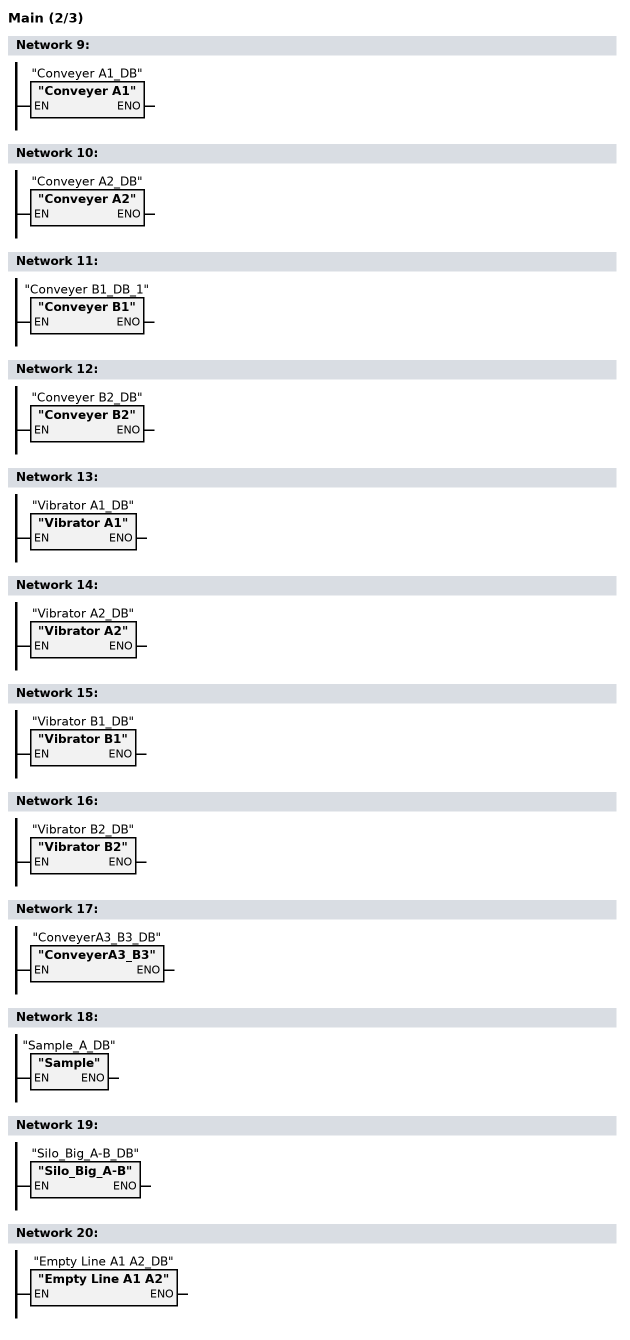
   RUNG wire#powerrail
      "Conveyer A1_DB"()
   END_RUNG
   // the same network as SCL:
   "Conveyer A1_DB"();   // "Conveyer A1"
END_REGION

REGION Network 10
   RUNG wire#powerrail
      "Conveyer A2_DB"()
   END_RUNG
   // the same network as SCL:
   "Conveyer A2_DB"();   // "Conveyer A2"
END_REGION

REGION Network 11
   RUNG wire#powerrail
      "Conveyer B1_DB_1"()
   END_RUNG
   // the same network as SCL:
   "Conveyer B1_DB_1"();   // "Conveyer B1"
END_REGION

REGION Network 12
   RUNG wire#powerrail
      "Conveyer B2_DB"()
   END_RUNG
   // the same network as SCL:
   "Conveyer B2_DB"();   // "Conveyer B2"
END_REGION

REGION Network 13
   RUNG wire#powerrail
      "Vibrator A1_DB"()
   END_RUNG
   // the same network as SCL:
   "Vibrator A1_DB"();   // "Vibrator A1"
END_REGION

REGION Network 14
   RUNG wire#powerrail
      "Vibrator A2_DB"()
   END_RUNG
   // the same network as SCL:
   "Vibrator A2_DB"();   // "Vibrator A2"
END_REGION

REGION Network 15
   RUNG wire#powerrail
      "Vibrator B1_DB"()
   END_RUNG
   // the same network as SCL:
   "Vibrator B1_DB"();   // "Vibrator B1"
END_REGION

REGION Network 16
   RUNG wire#powerrail
      "Vibrator B2_DB"()
   END_RUNG
   // the same network as SCL:
   "Vibrator B2_DB"();   // "Vibrator B2"
END_REGION

REGION Network 17
   RUNG wire#powerrail
      "ConveyerA3_B3_DB"()
   END_RUNG
   // the same network as SCL:
   "ConveyerA3_B3_DB"();   // "ConveyerA3_B3"
END_REGION

REGION Network 18
   RUNG wire#powerrail
      "Sample_A_DB"()
   END_RUNG
   // the same network as SCL:
   "Sample_A_DB"();   // "Sample"
END_REGION

REGION Network 19
   RUNG wire#powerrail
      "Silo_Big_A-B_DB"()
   END_RUNG
   // the same network as SCL:
   "Silo_Big_A-B_DB"();   // "Silo_Big_A-B"
END_REGION

REGION Network 20
   RUNG wire#powerrail
      "Empty Line A1 A2_DB"()
   END_RUNG
   // the same network as SCL:
   "Empty Line A1 A2_DB"();   // "Empty Line A1 A2"
END_REGION

REGION Network 21
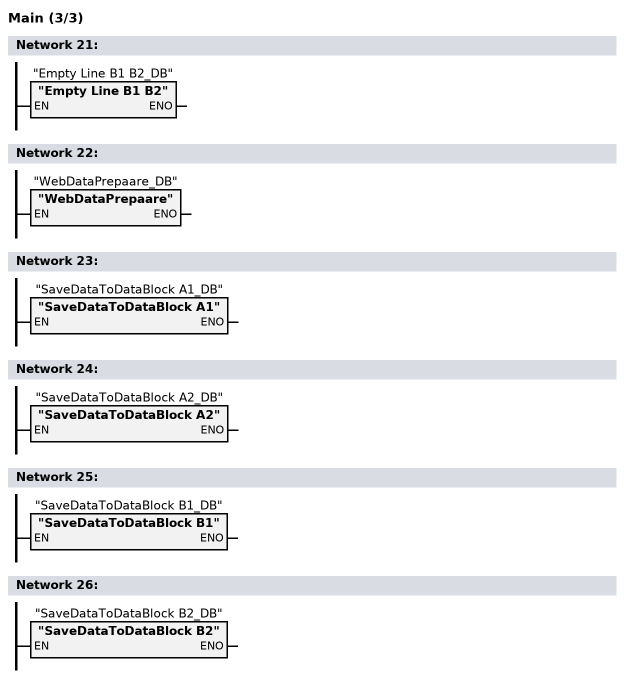
   RUNG wire#powerrail
      "Empty Line B1 B2_DB"()
   END_RUNG
   // the same network as SCL:
   "Empty Line B1 B2_DB"();   // "Empty Line B1 B2"
END_REGION

REGION Network 22
   RUNG wire#powerrail
      "WebDataPrepaare_DB"()
   END_RUNG
   // the same network as SCL:
   "WebDataPrepaare_DB"();   // "WebDataPrepaare"
END_REGION

REGION Network 23
   RUNG wire#powerrail
      "SaveDataToDataBlock A1_DB"()
   END_RUNG
   // the same network as SCL:
   "SaveDataToDataBlock A1_DB"();   // "SaveDataToDataBlock A1"
END_REGION

REGION Network 24
   RUNG wire#powerrail
      "SaveDataToDataBlock A2_DB"()
   END_RUNG
   // the same network as SCL:
   "SaveDataToDataBlock A2_DB"();   // "SaveDataToDataBlock A2"
END_REGION

REGION Network 25
   RUNG wire#powerrail
      "SaveDataToDataBlock B1_DB"()
   END_RUNG
   // the same network as SCL:
   "SaveDataToDataBlock B1_DB"();   // "SaveDataToDataBlock B1"
END_REGION

REGION Network 26
   RUNG wire#powerrail
      "SaveDataToDataBlock B2_DB"()
   END_RUNG
   // the same network as SCL:
   "SaveDataToDataBlock B2_DB"();   // "SaveDataToDataBlock B2"
END_REGION
END_ORGANIZATION_BLOCK

// ===== PLC "PLC_Lines_C"  CPU 1212C AC/DC/Rly =====

VAR_GLOBAL   // PLC tag table "Default tag table"
   "Tag_4" AT %MW114 : Word;
   "Tag_5" AT %M118.0 : Bool;
   "Tag_6" AT %M118.1 : Bool;
   "Tag_7" AT %M118.2 : Bool;
   "Tag_8" AT %MW120 : Word;
   "Tag_9" AT %MW122 : Word;
   "Tag_1" AT %M251.0 : Bool;
   "C2_Start_Conveyer" AT %M161.1 : Bool;
   "Tag_3" AT %M1000.0 : Bool;
   "Tag_10" AT %M1200.0 : Bool;
   "Vibrator_C1_On" AT %M151.4 : Bool;
   "Tag_11" AT %M151.5 : Bool;
   "Tag_2" AT %M123.2 : Bool;
   "Vibrator_C2_On" AT %M161.4 : Bool;
   "Tag_12" AT %M160.6 : Bool;
   "Conveyer_C2_On" AT %M160.3 : Bool;
   "Tag_13" AT %M161.5 : Bool;
   "Tag_14" AT %M151.7 : Bool;
   "Conveyer_C1_OneShut" AT %M151.3 : Bool;
   "Conveyer_C2_OneShut" AT %M161.3 : Bool;
   "Silo C Big" AT %Q3.6 : Bool;
   "Silo_C_Big_Start_Toggle" AT %M190.0 : Bool;
   "TriggerStartToggleMemory" AT %M152.0 : Bool;
   "TriggerC1ToggleStop" AT %M152.1 : Bool;
   "Conveyor_C1_Empty_line" AT %M152.2 : Bool;
   "Line_C2_Conveyer_Timer" AT %M162.0 : Bool;
   "TriggerStartToggleMemoryC2" AT %M162.1 : Bool;
   "TriggerStopToggleMemoryC21" AT %M162.2 : Bool;
   "Conveyor_C2_Empty_line" AT %M162.3 : Bool;
   "Silo_C_Not_Start_Timer" AT %M180.0 : Bool;
   "SiloCToggleStart" AT %M180.1 : Bool;
   "Tag_15" AT %MD210 : DInt;
   "Tag_16" AT %MD240 : DInt;
   "Tag_17" AT %M500.1 : Bool;
   "Tag_18" AT %M500.2 : Bool;
   "Tag_24" AT %MW502 : Word;
   "Tag_26" AT %M504.0 : Bool;
   "Tag_27" AT %M504.1 : Bool;
   "Tag_28" AT %M504.2 : Bool;
   "Tag_29" AT %MW506 : Word;
   "Tag_30" AT %MW508 : Word;
   "Tag_31" AT %MW510 : Word;
   "Tag_32" AT %M504.7 : Bool;
END_VAR

VAR_GLOBAL   // PLC tag table "InputOutput"
   "Emergency_C" AT %I0.6 : Bool;   // OK
   "Low_Silo_C1" AT %I0.2 : Bool;   // OK
   "Conveyer_C1" AT %Q0.2 : Bool;   // OK
   "Conveyer_C2" AT %Q0.3 : Bool;   // OK
   "Rel Out Vibrator C1" AT %Q0.0 : Bool;
   "Rel Out Vibrator C2" AT %Q0.1 : Bool;
   "Rel Out Alarm C1" AT %Q2.2 : Bool;
   "Rel Out Alarm C2" AT %Q2.3 : Bool;
   "Pneumatic_C1" AT %Q0.4 : Bool;   // OK
   "Pneumatic_C2" AT %Q0.5 : Bool;   // OK
   "Rel Out Conveyer C" AT %Q2.4 : Bool;
   "Rel Out Silo C Stop" AT %Q2.5 : Bool;
   "Rel Out Silo C Start" AT %Q2.6 : Bool;
   "Low_Silo_C2" AT %I0.0 : Bool;   // OK
   "HIgh_Silo_C1" AT %I0.3 : Bool;   // OK
   "Fault_C1" AT %I0.4 : Bool;   // OK
   "Fault_C2" AT %I0.5 : Bool;   // OK
   "High_Silo_C2" AT %I0.1 : Bool;   // OK
   "Start" AT %I1.1 : Bool;
   "Fault_C3" AT %I0.7 : Bool;   // OK
   "Conveyer_C3" AT %Q3.4 : Bool;   // OK
   "Light_C1" AT %Q2.0 : Bool;   // OK
   "Light_C2" AT %Q2.1 : Bool;   // OK
END_VAR

VAR_GLOBAL   // PLC tag table "SystemTag"
   "System_Byte" AT %MB1 : Byte;
   "FirstScan" AT %M1.0 : Bool;
   "DiagStatusUpdate" AT %M1.1 : Bool;
   "AlwaysTRUE" AT %M1.2 : Bool;
   "AlwaysFALSE" AT %M1.3 : Bool;
   "Clock_Byte" AT %MB0 : Byte;
   "Clock_10Hz" AT %M0.0 : Bool;
   "Clock_5Hz" AT %M0.1 : Bool;
   "Clock_2.5Hz" AT %M0.2 : Bool;
   "Clock_2Hz" AT %M0.3 : Bool;
   "Clock_1.25Hz" AT %M0.4 : Bool;
   "Clock_1Hz" AT %M0.5 : Bool;
   "Clock_0.625Hz" AT %M0.6 : Bool;
   "Clock_0.5Hz" AT %M0.7 : Bool;
   "DoneModbusCommon" AT %M110.0 : Bool;
   "ErrorModbusCommon" AT %M110.1 : Bool;
   "ModbusCommonStatus" AT %MW112 : Word;
END_VAR

VAR_GLOBAL   // PLC tag table "LineC1Tags"
   "Line_C1_Start_Consent" AT %M150.0 : Bool;
   "Line_C1_Run_Consent" AT %M150.1 : Bool;
   "Line_C1_Conveyer_Timer" AT %M150.2 : Bool;
   "Conveyer_C1_On" AT %M150.3 : Bool;
   "Conveyer_C1_Off" AT %M150.4 : Bool;
   "Line_C1_Light" AT %M151.0 : Bool;
   "Start_C1_Toggle" AT %M150.5 : Bool;
   "StartTriggerRisingTrigger" AT %M150.6 : Bool;
   "Conveyer_C1_Start_Consent" AT %M250.0 : Bool;
   "Conveyer_C1_Run_Consent" AT %M250.1 : Bool;
   "Silo_C_Start" AT %M300.0 : Bool;
   "C1_Sample_Triger" AT %M150.7 : Bool;
   "C1_Start_Conveyer" AT %M151.1 : Bool;
END_VAR

VAR_GLOBAL   // PLC tag table "LineC2Tags"
   "Line_C2_Start_Consent" AT %M160.0 : Bool;
   "Line_C2_Run_Consent" AT %M160.1 : Bool;
   "Line_C2_Vibrator_Timer" AT %M160.2 : Bool;
   "Conveyer_C2_Off" AT %M160.4 : Bool;
   "Conveyer_C2_Start_Consent" AT %M260.0 : Bool;
   "Conveyer_C2_Run_Consent" AT %M260.1 : Bool;
   "Start_C2_Toggle" AT %M160.5 : Bool;
   "C2_Sample_Triger" AT %M160.7 : Bool;
END_VAR

TYPE "tIMEDATATYPE"
   STRUCT
      HOUR : String;
      MINUTE : String;
      DAY : String;
      MONTH : String;
      YEAR : String;
   END_STRUCT;
END_TYPE

DATA_BLOCK "ModbusDataSendToFeeders"   // DB7
{ S7_Optimized_Access := 'FALSE' }
VERSION : 0.1
   VAR
      dataforsend : Array[0..3] of Int;
   END_VAR
BEGIN
   dataforsend[0] := 0;
   dataforsend[1] := 0;
   dataforsend[2] := 0;
   dataforsend[3] := 0;
END_DATA_BLOCK

DATA_BLOCK "Clock"   // DB9
{ S7_Optimized_Access := 'TRUE' }
VERSION : 0.1
   VAR
      "time" : DTL;
   END_VAR
BEGIN
END_DATA_BLOCK

DATA_BLOCK "Conveyer C1_DB"   // DB16
{ S7_Optimized_Access := 'TRUE' }
VERSION : 0.1
// stored: InstanceOfName Conveyer C1
"Conveyer C1"
BEGIN
END_DATA_BLOCK

DATA_BLOCK "Web_Send"   // DB23
{ S7_Optimized_Access := 'TRUE' }
VERSION : 0.1
   VAR
      C1_Scenario_Type : Int := 2;
      C2_Scenario_Type : Int := 1;
      B1_Scenario_Type : Int := 1;
      B2_Scenario_Type : Int := 1;
      C_Emergency : Bool;
      B_Emergency : Bool;
      C1_Fault : Bool;
      C2_Fault : Bool;
      B1_Fault : Bool;
      B2_Fault : Bool;
      C3_Fault : Bool;
      B3_Fault : Bool;
      C1_Silo_Low : Bool;
      C2_Silo_Low : Bool;
      B1_Silo_Low : Bool;
      B2_Silo_Low : Bool;
      C1_Conveyer : Bool;
      C2_Conveyer : Bool;
      B1_Conveyer : Bool;
      B2_Conveyer : Bool;
      C3_Conveyor : Bool;
      B3_Left_Conveyer : Bool;
      C1_Silo_High : Bool;
      C2_Silo_High : Bool;
      B1_Silo_High : Bool;
      B2_Silo_High : Bool;
      C1_Sample : Bool;
      C2_Sample : Bool;
      B1_Sample : Bool;
      B2_Sample : Bool;
      C1_Running_Duration : Time;
      C1_Pause_Duration : Time;
      C1_Feeder_Vibration_Intensity : Int;
      C1_Ruuning_Online : Time;
      C1_Pause_Online : Time;
      C1_Sample_Interval : Time;
      C1_Sample_Duration : Time;
      C1_Sample_Online : Time;
      C1_Enable : Bool;
      C1_Start : Bool;
      C1_Big_Silo : Bool;
      B1_Running_Duration : Time;
      B1_Pause_Duration : Time;
      B1_Feeder_Vibration_Intensity : Int;
      B1_Ruuning_Online : Time;
      B1_Pause_Online : Time;
      B1_Sample_Interval : Time;
      B1_Sample_Duration : Time;
      B1_Sample_Online : Time;
      B1_Enable : Bool;
      B1_Start : Bool;
      B1_Big_Silo : Bool;
      C2_Running_Duration : Time;
      C2_Pause_Duration : Time;
      C2_Feeder_Vibration_Intensity : Int;
      C2_Ruuning_Online : Time;
      C2_Pause_Online : Time;
      C2_Sample_Interval : Time;
      C2_Sample_Duration : Time;
      C2_Sample_Online : Time;
      C2_Enable : Bool;
      C2_Start : Bool;
      C2_Big_Silo : Bool;
      B2_Running_Duration : Time;
      B2_Pause_Duration : Time;
      B2_Feeder_Vibration_Intensity : Int;
      B2_Ruuning_Online : Time;
      B2_Pause_Online : Time;
      B2_Sample_Interval : Time;
      B2_Sample_Duration : Time;
      B2_Sample_Online : Time;
      B2_Enable : Bool;
      B2_Start : Bool;
      B2_Big_Silo : Bool;
      C1_Manual : Bool;
      C2_Manual : Bool;
      B1_Manual : Bool;
      B2_Manual : Bool;
      C1_Feeder : Bool;
      C2_Feeder : Bool;
      B1_Feeder : Bool;
      B2_Feeder : Bool;
      C1_Duration_Big_Silo_Stop_Time : Time;
      C2_Duration_Big_Silo_Stop_Time : Time;
      B1_Duration_Big_Silo_Stop_Time : Time;
      B2_Duration_Big_Silo_Stop_Time : Time;
      C1_Empty_Line_Time : Time;
      C2_Empty_Line_Time : Time;
      B1_Empty_Line_Time : Time;
      B2_Empty_Line_Time : Time;
      C1_Feeder_Delay_After_Start_Time : Time;
      C2_Feeder_Delay_After_Start_Time : Time;
      B1_Feeder_Delay_After_Start_Time : Time;
      B2_Feeder_Delay_After_Start_Time : Time;
      C1_Feeder_Delay_Before_Stop_Time : Time;
      C2_Feeder_Delay_Before_Stop_Time : Time;
      B1_Feeder_Delay_Before_Stop_Time : Time;
      B2_Feeder_Delay_Before_Stop_Time : Time;
      C1_Feeder_Delay_Time : Time;
      C1_Feeder_Delay_Time_1 : Time;
      C1_Feeder_Delay_Time_2 : Time;
      C1_Feeder_Delay_Time_3 : Time;
      B3_Conveyor : Bool;
   END_VAR
BEGIN
END_DATA_BLOCK

DATA_BLOCK "Conveyer C2_DB"   // DB24
{ S7_Optimized_Access := 'TRUE' }
VERSION : 0.1
// stored: InstanceOfName Conveyer C2
"Conveyer C2"
BEGIN
END_DATA_BLOCK

DATA_BLOCK "Vibrator C1_DB"   // DB25
{ S7_Optimized_Access := 'TRUE' }
VERSION : 0.1
// stored: InstanceOfName Vibrator C1
"Vibrator C1"
BEGIN
END_DATA_BLOCK

DATA_BLOCK "Vibrator C2_DB"   // DB26
{ S7_Optimized_Access := 'TRUE' }
VERSION : 0.1
// stored: InstanceOfName Vibrator C2
"Vibrator C2"
BEGIN
END_DATA_BLOCK

DATA_BLOCK "ConveyerC3_DB"   // DB35
{ S7_Optimized_Access := 'TRUE' }
VERSION : 0.1
// stored: InstanceOfName ConveyerC3
"ConveyerC3"
BEGIN
END_DATA_BLOCK

DATA_BLOCK "Sample_C_DB"   // DB36
{ S7_Optimized_Access := 'TRUE' }
VERSION : 0.1
// stored: InstanceOfName Sample_C
"Sample_C"
BEGIN
END_DATA_BLOCK

DATA_BLOCK "Silo_Big_C_DB"   // DB37
{ S7_Optimized_Access := 'TRUE' }
VERSION : 0.1
// stored: InstanceOfName Silo_Big_C
"Silo_Big_C"
BEGIN
END_DATA_BLOCK

DATA_BLOCK "Empty Line C1_DB"   // DB38
{ S7_Optimized_Access := 'TRUE' }
VERSION : 0.1
// stored: InstanceOfName Empty Line C1
"Empty Line C1"
BEGIN
END_DATA_BLOCK

DATA_BLOCK "Web_Recieve"   // DB45
{ S7_Optimized_Access := 'TRUE' }
VERSION : 0.1
   VAR
      Scenario_Type : Int;   // 1 2 3 4 5 A B C D E F
      Line_C1_Start : Bool;
      Line_C1_Enable : Bool := 0;
      Line_C2_Start : Bool;
      Line_C2_Enable : Bool;
      Line_C1_Conveyer_on_Time : Time := T#8S_400MS;
      Line_C1_Conveyer_off_Time : Time := T#30s;
      Line_C1_Sampling_Time : Time := T#2M;
      Line_C1_Sampling_OpenTime : Time := T#9S_500MS;
      Line_C2_Conveyer_on_Time : Time := T#8S_400MS;
      Line_C2_Conveyer_off_Time : Time := T#30s;
      Line_C2_Sampling_Time : Time := T#2M;
      Line_C2_Sampling_OpenTime : Time := T#9S_500MS;
      Line_C1_Feeder_Intensity : Int;
      Line_C2_Feeder_Intensity : Int;
      Line_C1_Feeder_DelayTime : Time;
      Line_C2_Feeder_DelayTime : Time;
      Line_C1_Enable_Manual : Bool;
      Line_C2_Enable_Manual : Bool;
      Line_C1_Conveyor_Start_Manual : Bool;
      Line_C2_Conveyor_Start_Manual : Bool;
      Line_C1_Big_Silo_Start_Manual : Bool;
      Line_C2_Big_Silo_Start_Manual : Bool;
      Line_C1_Below_Conveyor_Start_Manual : Bool;
      Line_C2_Below_Conveyor_Start_Manual : Bool;
      Line_C1_Feeder_Start_Manual : Bool;
      Line_C2_Feeder_Start_Manual : Bool;
      Line_B1_Feeder_Start_Manual : Bool;
      Line_B2_Feeder_Start_Manual : Bool;
      Line_C1_Sample_Start_Manual : Bool;
      Line_C2_Sample_Start_Manual : Bool;
      Line_B1_Sample_Start_Manual : Bool;
      Line_B2_Sample_Start_Manual : Bool;
      Line_C1_Feeder_Delay_Before_Stop_Time : Time;
      Line_B1_Feeder_Delay_Before_Stop_Time : Time;
      Line_C2_Feeder_Delay_Before_Stop_Time : Time;
      Line_B2_Feeder_Delay_Before_Stop_Time : Time;
      Line_C1_Empty_Line_Time : Time;
      Line_C2_Empty_Line_Time : Time;
      Line_B1_Empty_Line_Time : Time;
      Line_B2_Empty_Line_Time : Time;
      Line_C1_Big_Silo_Delay_Start : Time;
      Line_C2_Big_Silo_Delay_Start : Time;
      Line_B1_Big_Silo_Delay_Start : Time;
      Line_B2_Big_Silo_Delay_Start : Time;
      Line_C1_Empty_Line : Bool;
      Line_C2_Empty_Line : Bool;
      Line_B1_Empty_Line : Bool;
      Line_B2_Empty_Line : Bool;
      Line_C1_Feeder_Delay_After_Start_Time : Time;
      Line_C2_Feeder_Delay_After_Start_Time : Time;
      Line_B1_Feeder_Delay_After_Start_Time : Time;
      Line_B2_Feeder_Delay_After_Start_Time : Time;
   END_VAR
BEGIN
END_DATA_BLOCK

DATA_BLOCK "WebDataPrepaare_DB"   // DB49
{ S7_Optimized_Access := 'TRUE' }
VERSION : 0.1
// stored: InstanceOfName WebDataPrepaare
"WebDataPrepaare"
BEGIN
END_DATA_BLOCK

// folder: System blocks/Program resources

DATA_BLOCK "Timer_Before_On_Sample_C2"   // DB1
{ S7_Optimized_Access := 'TRUE' }
AUTHOR : Simatic
FAMILY : IEC
NAME : IEC_TMR
VERSION : 1.0
// stored: InstanceOfName IEC_TIMER
"IEC_TIMER"
BEGIN
END_DATA_BLOCK

DATA_BLOCK "Timer_C1_Empty_Line_DB"   // DB5
{ S7_Optimized_Access := 'TRUE' }
AUTHOR : Simatic
FAMILY : IEC
NAME : IEC_TMR
VERSION : 1.0
// stored: InstanceOfName IEC_TIMER
"IEC_TIMER"
BEGIN
END_DATA_BLOCK

DATA_BLOCK "Timer_C2_Empty_Line_DB"   // DB6
{ S7_Optimized_Access := 'TRUE' }
AUTHOR : Simatic
FAMILY : IEC
NAME : IEC_TMR
VERSION : 1.0
// stored: InstanceOfName IEC_TIMER
"IEC_TIMER"
BEGIN
END_DATA_BLOCK

DATA_BLOCK "Timer_Sample_Open_Time_C2"   // DB8
{ S7_Optimized_Access := 'TRUE' }
AUTHOR : Simatic
FAMILY : IEC
NAME : IEC_TMR
VERSION : 1.0
// stored: InstanceOfName IEC_TIMER
"IEC_TIMER"
BEGIN
END_DATA_BLOCK

DATA_BLOCK "Timer_Silo_Big_C_Off_Time"   // DB10
{ S7_Optimized_Access := 'TRUE' }
AUTHOR : Simatic
FAMILY : IEC
NAME : IEC_TMR
VERSION : 1.0
// stored: InstanceOfName IEC_TIMER
"IEC_TIMER"
BEGIN
END_DATA_BLOCK

DATA_BLOCK "C1_Feeder_On_Delay_Timer"   // DB11
{ S7_Optimized_Access := 'TRUE' }
AUTHOR : Simatic
FAMILY : IEC
NAME : IEC_TMR
VERSION : 1.0
// stored: InstanceOfName IEC_TIMER
"IEC_TIMER"
BEGIN
END_DATA_BLOCK

DATA_BLOCK "C2_Feeder_On_Delay_Timer"   // DB14
{ S7_Optimized_Access := 'TRUE' }
AUTHOR : Simatic
FAMILY : IEC
NAME : IEC_TMR
VERSION : 1.0
// stored: InstanceOfName IEC_TIMER
"IEC_TIMER"
BEGIN
END_DATA_BLOCK

DATA_BLOCK "IEC_Counter_0_DB"   // DB15
{ S7_Optimized_Access := 'TRUE' }
AUTHOR : Simatic
FAMILY : IEC
NAME : CNTR
VERSION : 1.0
// stored: InstanceOfName IEC_COUNTER
"IEC_COUNTER"
BEGIN
END_DATA_BLOCK

DATA_BLOCK "Timer_Off_C1_Conveyer"   // DB27
{ S7_Optimized_Access := 'TRUE' }
AUTHOR : Simatic
FAMILY : IEC
NAME : IEC_TMR
VERSION : 1.0
// stored: InstanceOfName IEC_TIMER
"IEC_TIMER"
BEGIN
END_DATA_BLOCK

DATA_BLOCK "Timer_On_C2_Conveyer"   // DB28
{ S7_Optimized_Access := 'TRUE' }
AUTHOR : Simatic
FAMILY : IEC
NAME : IEC_TMR
VERSION : 1.0
// stored: InstanceOfName IEC_TIMER
"IEC_TIMER"
BEGIN
END_DATA_BLOCK

DATA_BLOCK "Timer_Off_C2_Conveyer"   // DB29
{ S7_Optimized_Access := 'TRUE' }
AUTHOR : Simatic
FAMILY : IEC
NAME : IEC_TMR
VERSION : 1.0
// stored: InstanceOfName IEC_TIMER
"IEC_TIMER"
BEGIN
END_DATA_BLOCK

DATA_BLOCK "Timer_Before_On_Sample_C1"   // DB30
{ S7_Optimized_Access := 'TRUE' }
AUTHOR : Simatic
FAMILY : IEC
NAME : IEC_TMR
VERSION : 1.0
// stored: InstanceOfName IEC_TIMER
"IEC_TIMER"
BEGIN
END_DATA_BLOCK

DATA_BLOCK "Timer_Sample_Open_Time_C1"   // DB31
{ S7_Optimized_Access := 'TRUE' }
AUTHOR : Simatic
FAMILY : IEC
NAME : IEC_TMR
VERSION : 1.0
// stored: InstanceOfName IEC_TIMER
"IEC_TIMER"
BEGIN
END_DATA_BLOCK

DATA_BLOCK "Timer_On_C1_Conveyer"   // DB39
{ S7_Optimized_Access := 'TRUE' }
AUTHOR : Simatic
FAMILY : IEC
NAME : IEC_TMR
VERSION : 1.0
// stored: InstanceOfName IEC_TIMER
"IEC_TIMER"
BEGIN
END_DATA_BLOCK

// folder: (top level)

FUNCTION_BLOCK "Conveyer C1"   // FB1, LAD
{ S7_Optimized_Access := 'TRUE' }
VERSION : 0.1
   VAR_TEMP   // added for the SCL form of the ladder/FBD networks
      _w1 : Bool;
      _w2 : Bool;
   END_VAR
BEGIN

REGION Network 1: Start Consent line C1
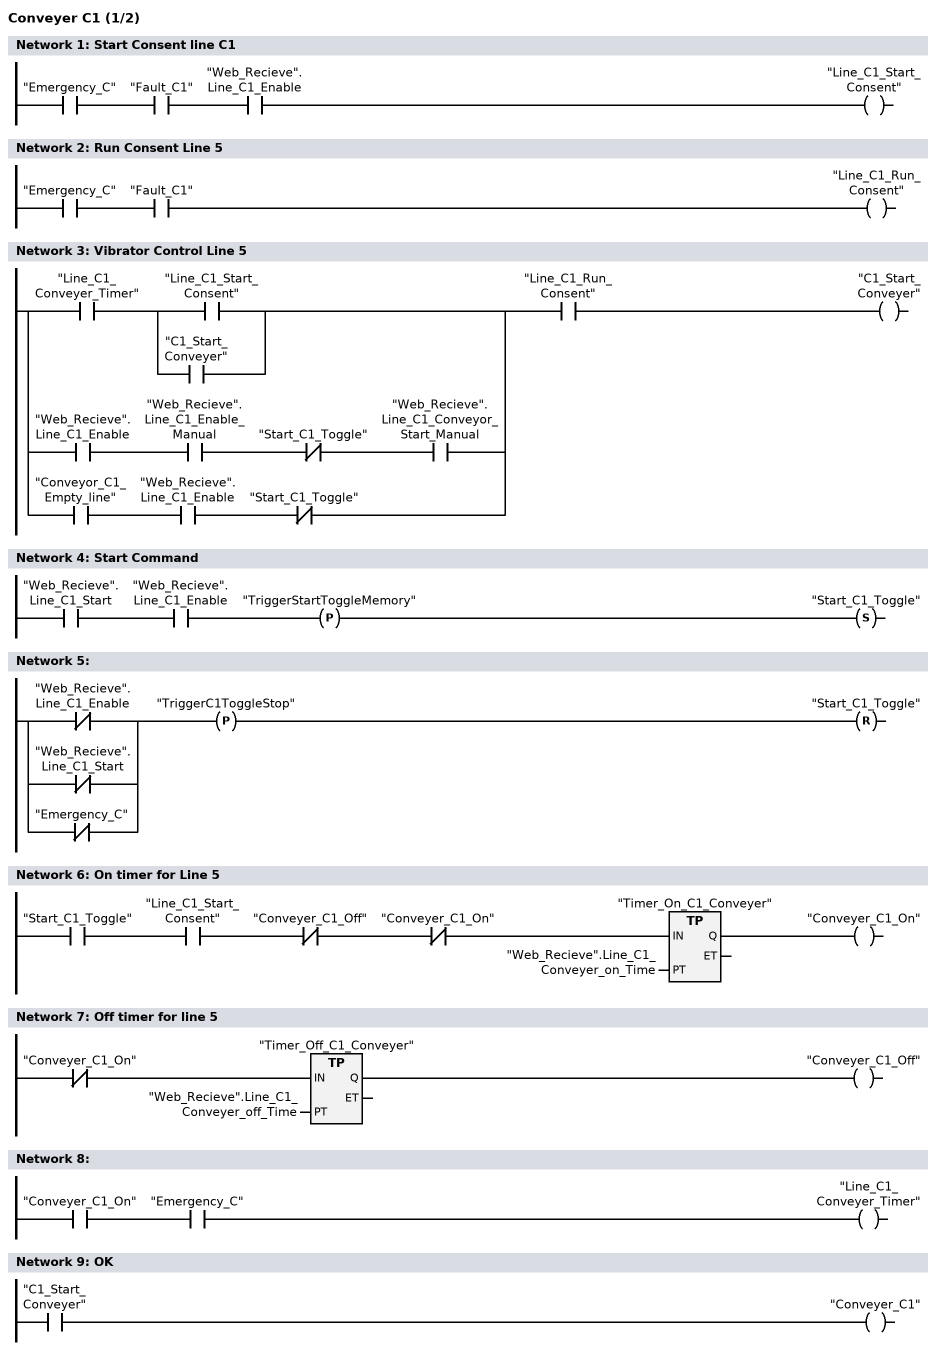
   RUNG wire#powerrail
      Contact( "Emergency_C" )
      Contact( "Fault_C1" )
      Contact( "Web_Recieve".Line_C1_Enable )
      Coil( "Line_C1_Start_Consent" )
   END_RUNG
   // the same network as SCL:
   "Line_C1_Start_Consent" := "Emergency_C" AND "Fault_C1" AND "Web_Recieve".Line_C1_Enable;
END_REGION

REGION Network 2: Run Consent Line 5
   RUNG wire#powerrail
      Contact( "Emergency_C" )
      Contact( "Fault_C1" )
      Coil( "Line_C1_Run_Consent" )
   END_RUNG
   // the same network as SCL:
   "Line_C1_Run_Consent" := "Emergency_C" AND "Fault_C1";
END_REGION

REGION Network 3: Vibrator Control Line 5
   RUNG wire#powerrail
      Contact( "Line_C1_Conveyer_Timer" )
      wire#w1
      Contact( "Line_C1_Start_Consent" )
      wire#w2
      Contact( "Line_C1_Run_Consent" )
      Coil( "C1_Start_Conveyer" )
   END_RUNG
   RUNG wire#w1
      Contact( "C1_Start_Conveyer" )
   END_RUNG wire#w2
   RUNG wire#powerrail
      Contact( "Web_Recieve".Line_C1_Enable )
      Contact( "Web_Recieve".Line_C1_Enable_Manual )
      I_Contact( "Start_C1_Toggle" )
      Contact( "Web_Recieve".Line_C1_Conveyor_Start_Manual )
   END_RUNG wire#w2
   RUNG wire#powerrail
      Contact( "Conveyor_C1_Empty_line" )
      Contact( "Web_Recieve".Line_C1_Enable )
      I_Contact( "Start_C1_Toggle" )
   END_RUNG wire#w2
   // the same network as SCL:
   "C1_Start_Conveyer" := (("Line_C1_Conveyer_Timer" AND ("Line_C1_Start_Consent" OR "C1_Start_Conveyer")) OR ("Web_Recieve".Line_C1_Enable AND "Web_Recieve".Line_C1_Enable_Manual AND NOT "Start_C1_Toggle" AND "Web_Recieve".Line_C1_Conveyor_Start_Manual) OR ("Conveyor_C1_Empty_line" AND "Web_Recieve".Line_C1_Enable AND NOT "Start_C1_Toggle")) AND "Line_C1_Run_Consent";
END_REGION

REGION Network 4: Start Command
   RUNG wire#powerrail
      Contact( "Web_Recieve".Line_C1_Start )
      Contact( "Web_Recieve".Line_C1_Enable )
      P_Trig( "TriggerStartToggleMemory" )
      S_Coil( "Start_C1_Toggle" )
   END_RUNG
   // the same network as SCL:
   #_w1 := "Web_Recieve".Line_C1_Start AND "Web_Recieve".Line_C1_Enable;
   #_w2 := #_w1 AND NOT "TriggerStartToggleMemory";   // rising edge
   "TriggerStartToggleMemory" := #_w1;
   IF #_w2 THEN "Start_C1_Toggle" := TRUE; END_IF;
END_REGION

REGION Network 5
   RUNG wire#powerrail
      I_Contact( "Web_Recieve".Line_C1_Enable )
      wire#w1
      P_Trig( "TriggerC1ToggleStop" )
      R_Coil( "Start_C1_Toggle" )
   END_RUNG
   RUNG wire#powerrail
      I_Contact( "Web_Recieve".Line_C1_Start )
   END_RUNG wire#w1
   RUNG wire#powerrail
      I_Contact( "Emergency_C" )
   END_RUNG wire#w1
   // the same network as SCL:
   #_w1 := NOT "Web_Recieve".Line_C1_Enable OR NOT "Web_Recieve".Line_C1_Start OR NOT "Emergency_C";
   #_w2 := #_w1 AND NOT "TriggerC1ToggleStop";   // rising edge
   "TriggerC1ToggleStop" := #_w1;
   IF #_w2 THEN "Start_C1_Toggle" := FALSE; END_IF;
END_REGION

REGION Network 6: On timer for Line 5
   "Timer_On_C1_Conveyer".TP(IN := "Start_C1_Toggle" AND "Line_C1_Start_Consent" AND NOT "Conveyer_C1_Off" AND NOT "Conveyer_C1_On",
                           PT := "Web_Recieve".Line_C1_Conveyer_on_Time);
   "Conveyer_C1_On" := "Timer_On_C1_Conveyer".Q;
END_REGION

REGION Network 7: Off timer for line 5
   "Timer_Off_C1_Conveyer".TP(IN := NOT "Conveyer_C1_On", PT := "Web_Recieve".Line_C1_Conveyer_off_Time);
   "Conveyer_C1_Off" := "Timer_Off_C1_Conveyer".Q;
END_REGION

REGION Network 8
   RUNG wire#powerrail
      Contact( "Conveyer_C1_On" )
      Contact( "Emergency_C" )
      Coil( "Line_C1_Conveyer_Timer" )
   END_RUNG
   // the same network as SCL:
   "Line_C1_Conveyer_Timer" := "Conveyer_C1_On" AND "Emergency_C";
END_REGION

REGION Network 9: OK
   RUNG wire#powerrail
      Contact( "C1_Start_Conveyer" )
      Coil( "Conveyer_C1" )
   END_RUNG
   // the same network as SCL:
   "Conveyer_C1" := "C1_Start_Conveyer";
END_REGION

REGION Network 10
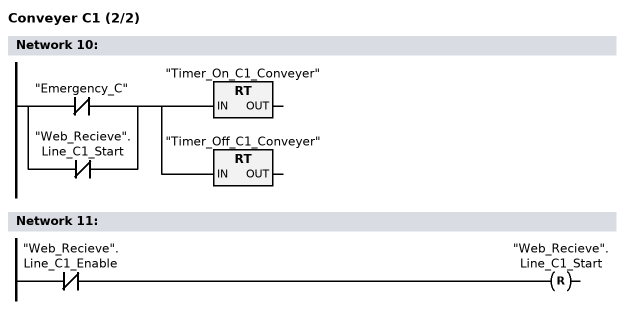
   RUNG wire#powerrail
      I_Contact( "Emergency_C" )
      wire#w1
      RT_Coil( "Timer_On_C1_Conveyer" )
   END_RUNG
   RUNG wire#powerrail
      I_Contact( "Web_Recieve".Line_C1_Start )
   END_RUNG wire#w1
   RUNG wire#w1
      RT_Coil( "Timer_Off_C1_Conveyer" )
   END_RUNG
   // the same network as SCL:
   #_w1 := NOT "Emergency_C" OR NOT "Web_Recieve".Line_C1_Start;
   IF #_w1 THEN
       RESET_TIMER("Timer_On_C1_Conveyer");
       RESET_TIMER("Timer_Off_C1_Conveyer");
   END_IF;
END_REGION

REGION Network 11
   RUNG wire#powerrail
      I_Contact( "Web_Recieve".Line_C1_Enable )
      R_Coil( "Web_Recieve".Line_C1_Start )
   END_RUNG
   // the same network as SCL:
   IF NOT "Web_Recieve".Line_C1_Enable THEN "Web_Recieve".Line_C1_Start := FALSE; END_IF;
END_REGION
END_FUNCTION_BLOCK

FUNCTION_BLOCK "Conveyer C2"   // FB2, LAD
{ S7_Optimized_Access := 'TRUE' }
VERSION : 0.1
   VAR_TEMP   // added for the SCL form of the ladder/FBD networks
      _w1 : Bool;
      _w2 : Bool;
   END_VAR
BEGIN

REGION Network 1: Start Consent line A1
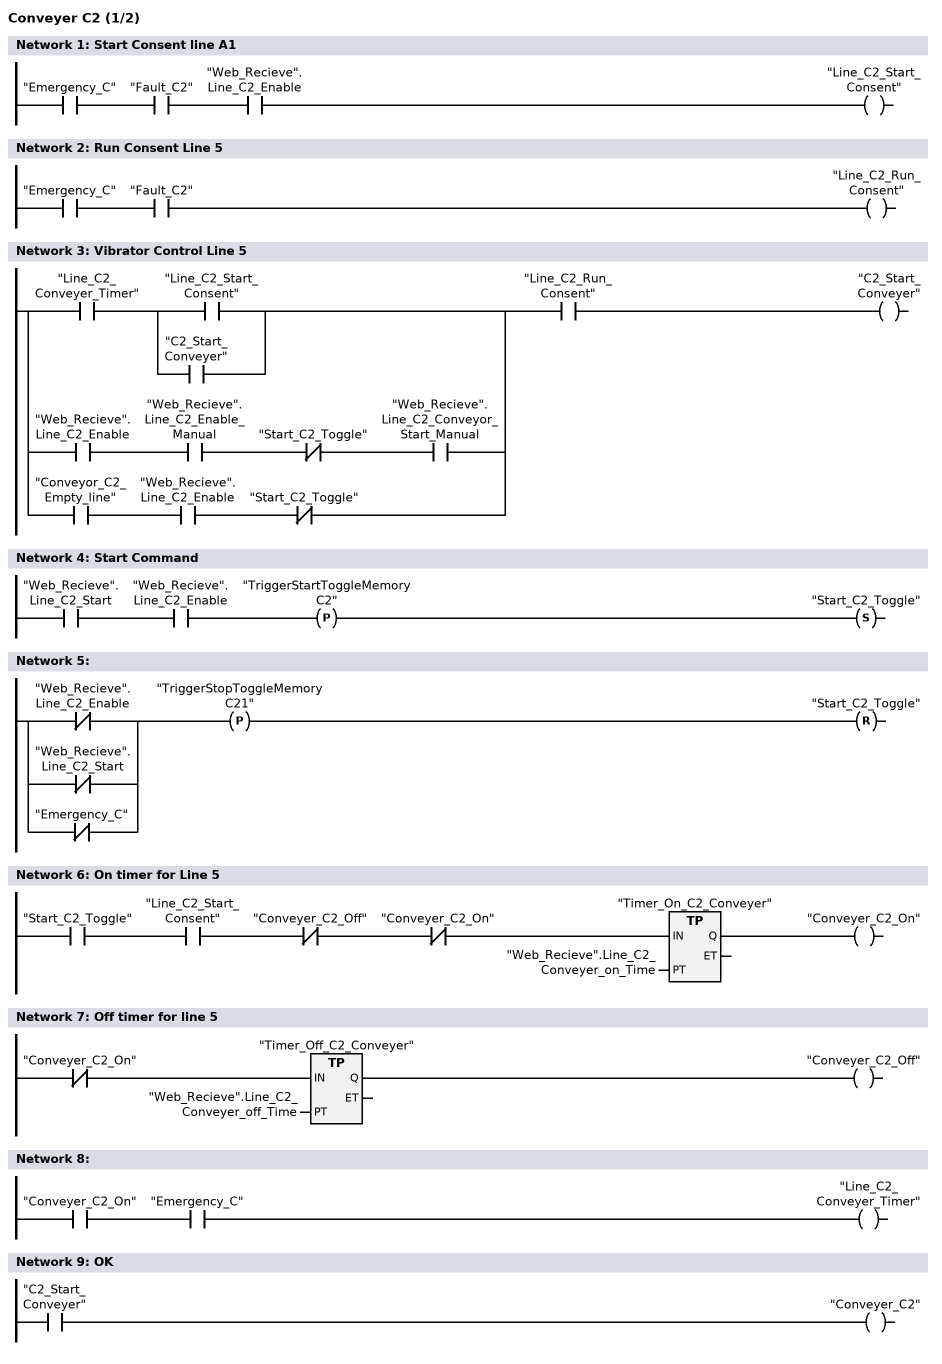
   RUNG wire#powerrail
      Contact( "Emergency_C" )
      Contact( "Fault_C2" )
      Contact( "Web_Recieve".Line_C2_Enable )
      Coil( "Line_C2_Start_Consent" )
   END_RUNG
   // the same network as SCL:
   "Line_C2_Start_Consent" := "Emergency_C" AND "Fault_C2" AND "Web_Recieve".Line_C2_Enable;
END_REGION

REGION Network 2: Run Consent Line 5
   RUNG wire#powerrail
      Contact( "Emergency_C" )
      Contact( "Fault_C2" )
      Coil( "Line_C2_Run_Consent" )
   END_RUNG
   // the same network as SCL:
   "Line_C2_Run_Consent" := "Emergency_C" AND "Fault_C2";
END_REGION

REGION Network 3: Vibrator Control Line 5
   RUNG wire#powerrail
      Contact( "Line_C2_Conveyer_Timer" )
      wire#w1
      Contact( "Line_C2_Start_Consent" )
      wire#w2
      Contact( "Line_C2_Run_Consent" )
      Coil( "C2_Start_Conveyer" )
   END_RUNG
   RUNG wire#w1
      Contact( "C2_Start_Conveyer" )
   END_RUNG wire#w2
   RUNG wire#powerrail
      Contact( "Web_Recieve".Line_C2_Enable )
      Contact( "Web_Recieve".Line_C2_Enable_Manual )
      I_Contact( "Start_C2_Toggle" )
      Contact( "Web_Recieve".Line_C2_Conveyor_Start_Manual )
   END_RUNG wire#w2
   RUNG wire#powerrail
      Contact( "Conveyor_C2_Empty_line" )
      Contact( "Web_Recieve".Line_C2_Enable )
      I_Contact( "Start_C2_Toggle" )
   END_RUNG wire#w2
   // the same network as SCL:
   "C2_Start_Conveyer" := (("Line_C2_Conveyer_Timer" AND ("Line_C2_Start_Consent" OR "C2_Start_Conveyer")) OR ("Web_Recieve".Line_C2_Enable AND "Web_Recieve".Line_C2_Enable_Manual AND NOT "Start_C2_Toggle" AND "Web_Recieve".Line_C2_Conveyor_Start_Manual) OR ("Conveyor_C2_Empty_line" AND "Web_Recieve".Line_C2_Enable AND NOT "Start_C2_Toggle")) AND "Line_C2_Run_Consent";
END_REGION

REGION Network 4: Start Command
   RUNG wire#powerrail
      Contact( "Web_Recieve".Line_C2_Start )
      Contact( "Web_Recieve".Line_C2_Enable )
      P_Trig( "TriggerStartToggleMemoryC2" )
      S_Coil( "Start_C2_Toggle" )
   END_RUNG
   // the same network as SCL:
   #_w1 := "Web_Recieve".Line_C2_Start AND "Web_Recieve".Line_C2_Enable;
   #_w2 := #_w1 AND NOT "TriggerStartToggleMemoryC2";   // rising edge
   "TriggerStartToggleMemoryC2" := #_w1;
   IF #_w2 THEN "Start_C2_Toggle" := TRUE; END_IF;
END_REGION

REGION Network 5
   RUNG wire#powerrail
      I_Contact( "Web_Recieve".Line_C2_Enable )
      wire#w1
      P_Trig( "TriggerStopToggleMemoryC21" )
      R_Coil( "Start_C2_Toggle" )
   END_RUNG
   RUNG wire#powerrail
      I_Contact( "Web_Recieve".Line_C2_Start )
   END_RUNG wire#w1
   RUNG wire#powerrail
      I_Contact( "Emergency_C" )
   END_RUNG wire#w1
   // the same network as SCL:
   #_w1 := NOT "Web_Recieve".Line_C2_Enable OR NOT "Web_Recieve".Line_C2_Start OR NOT "Emergency_C";
   #_w2 := #_w1 AND NOT "TriggerStopToggleMemoryC21";   // rising edge
   "TriggerStopToggleMemoryC21" := #_w1;
   IF #_w2 THEN "Start_C2_Toggle" := FALSE; END_IF;
END_REGION

REGION Network 6: On timer for Line 5
   "Timer_On_C2_Conveyer".TP(IN := "Start_C2_Toggle" AND "Line_C2_Start_Consent" AND NOT "Conveyer_C2_Off" AND NOT "Conveyer_C2_On",
                           PT := "Web_Recieve".Line_C2_Conveyer_on_Time);
   "Conveyer_C2_On" := "Timer_On_C2_Conveyer".Q;
END_REGION

REGION Network 7: Off timer for line 5
   "Timer_Off_C2_Conveyer".TP(IN := NOT "Conveyer_C2_On", PT := "Web_Recieve".Line_C2_Conveyer_off_Time);
   "Conveyer_C2_Off" := "Timer_Off_C2_Conveyer".Q;
END_REGION

REGION Network 8
   RUNG wire#powerrail
      Contact( "Conveyer_C2_On" )
      Contact( "Emergency_C" )
      Coil( "Line_C2_Conveyer_Timer" )
   END_RUNG
   // the same network as SCL:
   "Line_C2_Conveyer_Timer" := "Conveyer_C2_On" AND "Emergency_C";
END_REGION

REGION Network 9: OK
   RUNG wire#powerrail
      Contact( "C2_Start_Conveyer" )
      Coil( "Conveyer_C2" )
   END_RUNG
   // the same network as SCL:
   "Conveyer_C2" := "C2_Start_Conveyer";
END_REGION

REGION Network 10
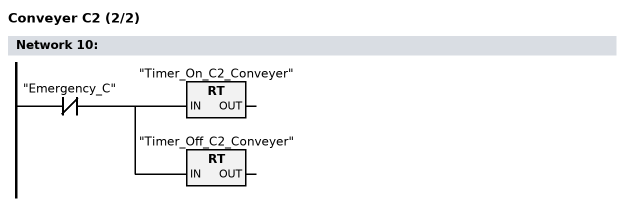
   RUNG wire#powerrail
      I_Contact( "Emergency_C" )
      wire#w1
      RT_Coil( "Timer_On_C2_Conveyer" )
   END_RUNG
   RUNG wire#w1
      RT_Coil( "Timer_Off_C2_Conveyer" )
   END_RUNG
   // the same network as SCL:
   IF NOT "Emergency_C" THEN
       RESET_TIMER("Timer_On_C2_Conveyer");
       RESET_TIMER("Timer_Off_C2_Conveyer");
   END_IF;
END_REGION
END_FUNCTION_BLOCK

FUNCTION_BLOCK "Vibrator C1"   // FB5, LAD
{ S7_Optimized_Access := 'TRUE' }
VERSION : 0.1
   VAR_TEMP
      RemainTime : DInt;
   END_VAR
BEGIN

REGION Network 1
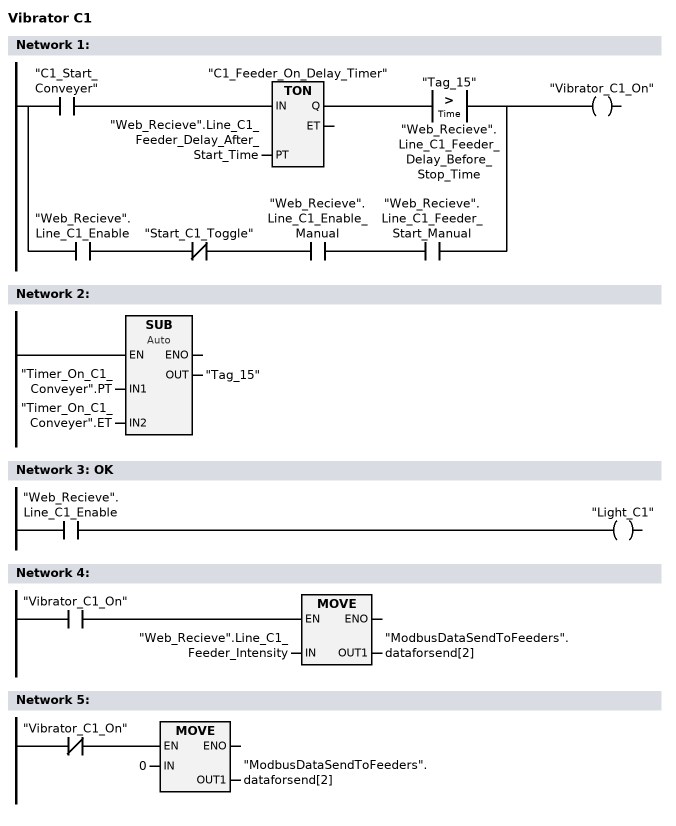
   "C1_Feeder_On_Delay_Timer".TON(IN := "C1_Start_Conveyer",
                           PT := "Web_Recieve".Line_C1_Feeder_Delay_After_Start_Time);
   "Vibrator_C1_On" := ("C1_Feeder_On_Delay_Timer".Q AND ("Tag_15" > "Web_Recieve".Line_C1_Feeder_Delay_Before_Stop_Time)) OR ("Web_Recieve".Line_C1_Enable AND NOT "Start_C1_Toggle" AND "Web_Recieve".Line_C1_Enable_Manual AND "Web_Recieve".Line_C1_Feeder_Start_Manual);
END_REGION

REGION Network 2
   RUNG wire#powerrail
      Sub(in1 := "Timer_On_C1_Conveyer".PT, in2 := "Timer_On_C1_Conveyer".ET, out => "Tag_15")
   END_RUNG
   // the same network as SCL:
   "Tag_15" := "Timer_On_C1_Conveyer".PT - "Timer_On_C1_Conveyer".ET;
END_REGION

REGION Network 3: OK
   RUNG wire#powerrail
      Contact( "Web_Recieve".Line_C1_Enable )
      Coil( "Light_C1" )
   END_RUNG
   // the same network as SCL:
   "Light_C1" := "Web_Recieve".Line_C1_Enable;
END_REGION

REGION Network 4
   RUNG wire#powerrail
      Contact( "Vibrator_C1_On" )
      Move(in := "Web_Recieve".Line_C1_Feeder_Intensity, out1 => "ModbusDataSendToFeeders".dataforsend[2])
   END_RUNG
   // the same network as SCL:
   IF "Vibrator_C1_On" THEN
       "ModbusDataSendToFeeders".dataforsend[2] := "Web_Recieve".Line_C1_Feeder_Intensity;
   END_IF;
END_REGION

REGION Network 5
   RUNG wire#powerrail
      I_Contact( "Vibrator_C1_On" )
      Move(in := 0, out1 => "ModbusDataSendToFeeders".dataforsend[2])
   END_RUNG
   // the same network as SCL:
   IF NOT "Vibrator_C1_On" THEN "ModbusDataSendToFeeders".dataforsend[2] := 0; END_IF;
END_REGION
END_FUNCTION_BLOCK

FUNCTION_BLOCK "Vibrator C2"   // FB6, LAD
{ S7_Optimized_Access := 'TRUE' }
VERSION : 0.1
BEGIN

REGION Network 1
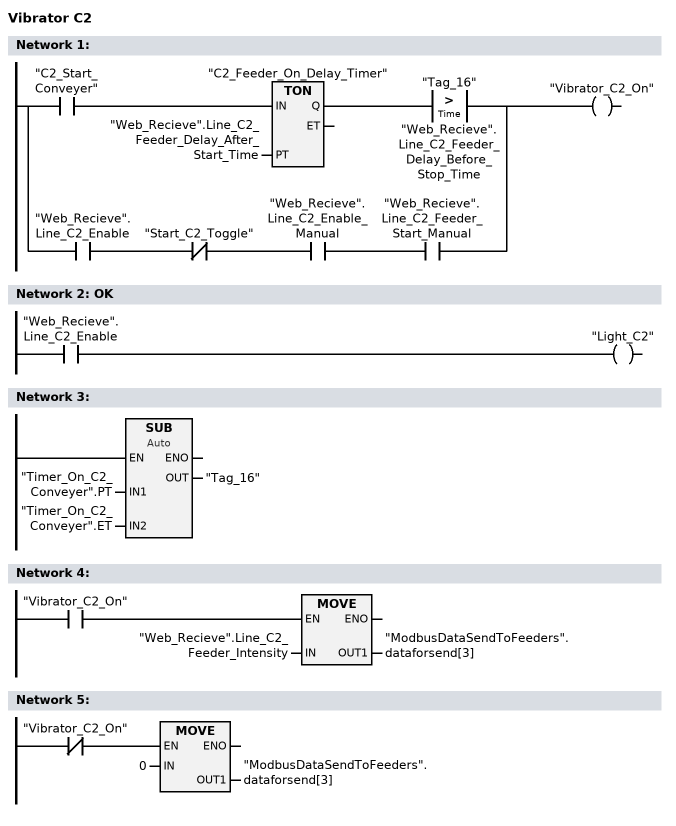
   "C2_Feeder_On_Delay_Timer".TON(IN := "C2_Start_Conveyer",
                           PT := "Web_Recieve".Line_C2_Feeder_Delay_After_Start_Time);
   "Vibrator_C2_On" := ("C2_Feeder_On_Delay_Timer".Q AND ("Tag_16" > "Web_Recieve".Line_C2_Feeder_Delay_Before_Stop_Time)) OR ("Web_Recieve".Line_C2_Enable AND NOT "Start_C2_Toggle" AND "Web_Recieve".Line_C2_Enable_Manual AND "Web_Recieve".Line_C2_Feeder_Start_Manual);
END_REGION

REGION Network 2: OK
   RUNG wire#powerrail
      Contact( "Web_Recieve".Line_C2_Enable )
      Coil( "Light_C2" )
   END_RUNG
   // the same network as SCL:
   "Light_C2" := "Web_Recieve".Line_C2_Enable;
END_REGION

REGION Network 3
   RUNG wire#powerrail
      Sub(in1 := "Timer_On_C2_Conveyer".PT, in2 := "Timer_On_C2_Conveyer".ET, out => "Tag_16")
   END_RUNG
   // the same network as SCL:
   "Tag_16" := "Timer_On_C2_Conveyer".PT - "Timer_On_C2_Conveyer".ET;
END_REGION

REGION Network 4
   RUNG wire#powerrail
      Contact( "Vibrator_C2_On" )
      Move(in := "Web_Recieve".Line_C2_Feeder_Intensity, out1 => "ModbusDataSendToFeeders".dataforsend[3])
   END_RUNG
   // the same network as SCL:
   IF "Vibrator_C2_On" THEN
       "ModbusDataSendToFeeders".dataforsend[3] := "Web_Recieve".Line_C2_Feeder_Intensity;
   END_IF;
END_REGION

REGION Network 5
   RUNG wire#powerrail
      I_Contact( "Vibrator_C2_On" )
      Move(in := 0, out1 => "ModbusDataSendToFeeders".dataforsend[3])
   END_RUNG
   // the same network as SCL:
   IF NOT "Vibrator_C2_On" THEN "ModbusDataSendToFeeders".dataforsend[3] := 0; END_IF;
END_REGION
END_FUNCTION_BLOCK

FUNCTION_BLOCK "ConveyerC3"   // FB9, LAD
{ S7_Optimized_Access := 'TRUE' }
VERSION : 0.1
BEGIN

REGION Network 1: OK